screen "0004_Mixinghead" 1280x800, template "Navigation"
   on GenerateScreen: SetBit("DB704_MH_Value_Read"); SetBit("DB614_MH_State_Read"); SetTag("Navigation_7", 4); "MH_TestshotVisibility"()
   Button "Button_17" at 118,142 size 357x253; TextOff 'Text'
      Visibility <- "MH_Control_Visibility"
   TextField "Text field_43" at 173,150 size 158x29; Text 'Temperature'
      Visibility <- "MH_Control_Visibility"
   TextField "Text field_44" at 124,193 size 72x25; Text 'Actual:'
      Visibility <- "MH_Control_Visibility"
   TextField "Text field_45" at 124,226 size 100x25; Text 'Set value:'
      Visibility <- "MH_Control_Visibility"
   TextField "Text field_46" at 124,259 size 201x25; Text 'Warning upper limit:'
      Visibility <- "MH_Control_Visibility"
   TextField "Text field_47" at 124,292 size 199x25; Text 'Warning lower limit:'
      Visibility <- "MH_Control_Visibility"
   TextField "Text field_48" at 124,325 size 170x25; Text 'Fault upper limit:'
      Visibility <- "MH_Control_Visibility"
   TextField "Text field_49" at 124,358 size 168x25; Text 'Fault lower limit:'
      Visibility <- "MH_Control_Visibility"
   IOField "I/O field_29" at 336,189 size 81x32; FormatPattern 999.9
      Visibility <- "MH_Control_Visibility"
      ProcessValue <- "Temp_Actual"
   IOField "I/O field_30" at 336,222 size 81x32; Authorization "Operate"; FormatPattern 999.9
      Visibility <- "MH_Control_Visibility"
      ProcessValue <- "Temp_SetValue"
   IOField "I/O field_31" at 336,255 size 81x32; Authorization "Operate"; FormatPattern 999.9
      Visibility <- "MH_Control_Visibility"
      ProcessValue <- "Temp_Warning_Upper_Limit"
   IOField "I/O field_32" at 336,288 size 81x32; Authorization "Operate"; FormatPattern 999.9
      Visibility <- "MH_Control_Visibility"
      ProcessValue <- "Temp_Warning_Llower_Limit"
   IOField "I/O field_33" at 336,321 size 81x32; Authorization "Operate"; FormatPattern 999.9
      Visibility <- "MH_Control_Visibility"
      ProcessValue <- "Temp_Fault_Upper_Limit"
   IOField "I/O field_34" at 336,354 size 81x32; Authorization "Operate"; FormatPattern 999.9
      Visibility <- "MH_Control_Visibility"
      ProcessValue <- "Temp_Fault_Lower_Limit"
   Button "Button_18" at 417,148 size 51x41; TextOff 'Text'; PictureOff "images (1)"
      on Press: SetTag("MH_Control_Visibility", 0)
      Visibility <- "MH_Control_Visibility"
   TextField "Text field_78" at 424,193 size 46x25; Text 'ºC'
      Visibility <- "MH_Control_Visibility"
   IOField "I/O field_50" at 317,150 size 84x30; FormatPattern ????????????????????
      Visibility <- "MH_Control_Visibility"
      ProcessValue <- "Temp_Name"
   TextField "Text field_42" at 424,226 size 46x25; Text 'ºC'
      Visibility <- "MH_Control_Visibility"
   TextField "Text field_50" at 424,259 size 46x25; Text 'Δ ºC'
      Visibility <- "MH_Control_Visibility"
   TextField "Text field_51" at 424,292 size 46x25; Text 'Δ ºC'
      Visibility <- "MH_Control_Visibility"
   TextField "Text field_52" at 424,325 size 46x25; Text 'Δ ºC'
      Visibility <- "MH_Control_Visibility"
   TextField "Text field_53" at 424,358 size 46x25; Text 'Δ ºC'
      Visibility <- "MH_Control_Visibility"
   Button "Button_7" at 117,142 size 357x253; TextOff 'Text'
      Visibility <- "MH_Control_Visibility"
   TextField "Text field_92" at 216,154 size 160x29; Text 'Inerting Data'
      Visibility <- "MH_Control_Visibility"
   TextField "Text field_93" at 123,189 size 118x25; Text 'Ready time:'
      Visibility <- "MH_Control_Visibility"
   TextField "Text field_94" at 123,217 size 188x25; Text 'Max. Inerting time:'
      Visibility <- "MH_Control_Visibility"
   TextField "Text field_95" at 123,245 size 198x25; Text 'Limit value inerting:'
      Visibility <- "MH_Control_Visibility"
   TextField "Text field_96" at 123,273 size 121x25; Text 'Start filling:'
      Visibility <- "MH_Control_Visibility"
   TextField "Text field_97" at 123,301 size 134x25; Text 'Filling factor:'
      Visibility <- "MH_Control_Visibility"
   TextField "Text field_98" at 123,329 size 122x25; Text 'Start offset:'
      Visibility <- "MH_Control_Visibility"
   IOField "I/O field_58" at 308,189 size 81x25; Authorization "Operate"; FormatPattern 99999
      Visibility <- "MH_Control_Visibility"
      ProcessValue <- "DB704_MH_Value_MH_Inerting{0}_Ready_Time_after_Inert"
   IOField "I/O field_59" at 308,217 size 81x25; Authorization "Operate"; FormatPattern 99999
      Visibility <- "MH_Control_Visibility"
      ProcessValue <- "DB704_MH_Value_MH_Inerting{0}_Max_Inerting_Time"
   IOField "I/O field_60" at 308,245 size 81x25; Authorization "User administration"; FormatPattern 9999.9
      Visibility <- "MH_Control_Visibility"
      ProcessValue <- "DB704_MH_Value_MH_Inerting{0}_Reference_Value_Inert"
   IOField "I/O field_61" at 308,273 size 81x25; Authorization "Operate"; FormatPattern 99999
      Visibility <- "MH_Control_Visibility"
      ProcessValue <- "DB704_MH_Value_MH_Inerting{0}_Foam_density"
   IOField "I/O field_62" at 308,301 size 81x25; Authorization "Operate"; FormatPattern 999.9
      Visibility <- "MH_Control_Visibility"
      ProcessValue <- "DB704_MH_Value_MH_Inerting{0}_Inerting_factor"
   IOField "I/O field_63" at 308,329 size 81x25; Authorization "Operate"; FormatPattern 999.9
      Visibility <- "MH_Control_Visibility"
      ProcessValue <- "DB704_MH_Value_MH_Inerting{0}_Start_Offset"
   Button "Button_9" at 416,148 size 51x41; TextOff 'Text'; PictureOff "images (1)"
      on Press: SetTag("MH_Control_Visibility", 0)
      Visibility <- "MH_Control_Visibility"
   IOField "I/O field_64" at 308,357 size 81x25; Authorization "Operate"; FormatPattern 999.9
      Visibility <- "MH_Control_Visibility"
      ProcessValue <- "DB704_MH_Value_MH_Inerting{0}_Leakage_Value"
   TextField "Text field_111" at 123,357 size 97x25; Text 'Min.level:'
      Visibility <- "MH_Control_Visibility"
   TextField "Text field_99" at 403,189 size 46x25; Text 's'
      Visibility <- "MH_Control_Visibility"
   TextField "Text field_100" at 403,217 size 46x25; Text 's'
      Visibility <- "MH_Control_Visibility"
   TextField "Text field_101" at 403,245 size 46x25; Text 'g'
      Visibility <- "MH_Control_Visibility"
   TextField "Text field_102" at 404,273 size 57x25; Text 'g/dm'
      Visibility <- "MH_Control_Visibility"
   TextField "Text field_103" at 452,269 size 36x18; Text '3'
      Visibility <- "MH_Control_Visibility"
   TextField "Text field_104" at 403,329 size 46x25; Text 'L'
      Visibility <- "MH_Control_Visibility"
   TextField "Text field_105" at 403,357 size 46x25; Text 'L'
      Visibility <- "MH_Control_Visibility"
   Button "Button_24" at 417,149 size 51x41; TextOff 'Text'; PictureOff "images (1)"
      on Press: SetTag("MH_Control_Visibility", 0)
      Visibility <- "MH_Control_Visibility"
   Button "Button_25" at 118,143 size 357x253; TextOff 'Text'
      Visibility <- "MH_Control_Visibility"
   TextField "Text field_137" at 249,155 size 96x29; Text 'Blowing'
      Visibility <- "MH_Control_Visibility"
   TextField "Text field_138" at 124,215 size 137x25; Text 'Blowing time:'
      Visibility <- "MH_Control_Visibility"
   TextField "Text field_139" at 124,248 size 237x25; Text 'Blowing time after shot:'
      Visibility <- "MH_Control_Visibility"
   IOField "I/O field_79" at 346,215 size 81x25; Authorization "Operate"; FormatPattern 99999
      Visibility <- "MH_Control_Visibility"
      ProcessValue <- "DB704_MH_Value_MH_Inerting{0}_Purge_time"
   IOField "I/O field_80" at 346,248 size 81x25; Authorization "Operate"; FormatPattern 99999
      Visibility <- "MH_Control_Visibility"
      ProcessValue <- "DB704_MH_Value_MH_Inerting{0}_Purge_after_Shot"
   Button "Button_26" at 417,149 size 51x41; TextOff 'Text'; PictureOff "images (1)"
      on Press: SetTag("MH_Control_Visibility", 0)
      Visibility <- "MH_Control_Visibility"
   TextField "Text field_145" at 442,215 size 46x25; Text 's'
      Visibility <- "MH_Control_Visibility"
   TextField "Text field_146" at 442,248 size 46x25; Text 's'
      Visibility <- "MH_Control_Visibility"
   Button "spare_2" at 335,709 size 36x32; TextOff 'Text'
      Visibility <- "DB704_MH_Value_Mixinghead{0}_MH_Connection{1}_WithNozzle"
   Button "spare_3" at 335,748 size 36x32; TextOff 'Text'
      Visibility <- "DB704_MH_Value_Mixinghead{0}_MH_Connection{1}_WithNozzle"
   Button "spare_1" at 335,670 size 36x32; TextOff 'Text'
      Visibility <- "DB704_MH_Value_Mixinghead{0}_MH_Connection{1}_WithNozzle"
   Button "spare_10" at 473,748 size 36x32; TextOff 'Text'
      Visibility <- "DB704_MH_Value_Mixinghead{0}_MH_Connection{2}_WithNozzle"
   Button "spare_9" at 473,709 size 36x32; TextOff 'Text'
      Visibility <- "DB704_MH_Value_Mixinghead{0}_MH_Connection{2}_WithNozzle"
   Button "spare_4" at 473,670 size 36x32; TextOff 'Text'
      Visibility <- "DB704_MH_Value_Mixinghead{0}_MH_Connection{2}_WithNozzle"
   Button "spare_5" at 611,670 size 36x32; TextOff 'Text'
      Visibility <- "DB704_MH_Value_Mixinghead{0}_MH_Connection{3}_WithNozzle"
   Button "spare_11" at 611,709 size 36x32; TextOff 'Text'
      Visibility <- "DB704_MH_Value_Mixinghead{0}_MH_Connection{3}_WithNozzle"
   Button "spare_12" at 611,748 size 36x32; TextOff 'Text'
      Visibility <- "DB704_MH_Value_Mixinghead{0}_MH_Connection{3}_WithNozzle"
   Button "spare_14" at 749,748 size 36x32; TextOff 'Text'
      Visibility <- "DB704_MH_Value_Mixinghead{0}_MH_Connection{4}_WithNozzle"
   Button "spare_13" at 749,709 size 36x32; TextOff 'Text'
      Visibility <- "DB704_MH_Value_Mixinghead{0}_MH_Connection{4}_WithNozzle"
   Button "spare_6" at 749,670 size 36x32; TextOff 'Text'
      Visibility <- "DB704_MH_Value_Mixinghead{0}_MH_Connection{4}_WithNozzle"
   Button "spare_7" at 887,670 size 36x32; TextOff 'Text'
      Visibility <- "DB704_MH_Value_Mixinghead{0}_MH_Connection{5}_WithNozzle"
   Button "spare_15" at 887,709 size 36x32; TextOff 'Text'
      Visibility <- "DB704_MH_Value_Mixinghead{0}_MH_Connection{5}_WithNozzle"
   Button "spare_16" at 887,748 size 36x32; TextOff 'Text'
      Visibility <- "DB704_MH_Value_Mixinghead{0}_MH_Connection{5}_WithNozzle"
   Button "spare_17" at 1025,709 size 36x32; TextOff 'Text'
      Visibility <- "DB704_MH_Value_Mixinghead{0}_MH_Connection{6}_WithNozzle"
   Button "spare_18" at 1025,748 size 36x32; TextOff 'Text'
      Visibility <- "DB704_MH_Value_Mixinghead{0}_MH_Connection{6}_WithNozzle"
   Button "spare_8" at 1025,670 size 36x32; TextOff 'Text'
      Visibility <- "DB704_MH_Value_Mixinghead{0}_MH_Connection{6}_WithNozzle"
   Rectangle "Rectangle_43" at 746,666 size 138x40
      Visibility <- "DB614_MH_State_MH_Status{0}_QPB_Values_selected"
   Rectangle "Rectangle_40" at 470,627 size 138x40
      Visibility <- "DB614_MH_State_MH_Status{0}_QPB_Values_selected"
   Rectangle "Rectangle_35" at 608,627 size 138x40
      Visibility <- "DB614_MH_State_MH_Status{0}_QPB_Values_selected"
   Rectangle "Rectangle_36" at 746,627 size 138x40
      Visibility <- "DB614_MH_State_MH_Status{0}_QPB_Values_selected"
   Rectangle "Rectangle_37" at 884,627 size 138x40
      Visibility <- "DB614_MH_State_MH_Status{0}_QPB_Values_selected"
   Rectangle "Rectangle_38" at 1022,627 size 138x40
      Visibility <- "DB614_MH_State_MH_Status{0}_QPB_Values_selected"
   Rectangle "Rectangle_41" at 470,666 size 138x40
      Visibility <- "DB614_MH_State_MH_Status{0}_QPB_Values_selected"
   Rectangle "Rectangle_42" at 608,666 size 138x40
      Visibility <- "DB614_MH_State_MH_Status{0}_QPB_Values_selected"
   Rectangle "Rectangle_44" at 884,666 size 138x40
      Visibility <- "DB614_MH_State_MH_Status{0}_QPB_Values_selected"
   Rectangle "Rectangle_45" at 1022,666 size 138x40
      Visibility <- "DB614_MH_State_MH_Status{0}_QPB_Values_selected"
   Rectangle "Rectangle_46" at 470,705 size 138x40
      Visibility <- "DB614_MH_State_MH_Status{0}_QPB_Values_selected"
   Rectangle "Rectangle_47" at 608,705 size 138x40
      Visibility <- "DB614_MH_State_MH_Status{0}_QPB_Values_selected"
   Rectangle "Rectangle_48" at 746,705 size 138x40
      Visibility <- "DB614_MH_State_MH_Status{0}_QPB_Values_selected"
   Rectangle "Rectangle_49" at 884,705 size 138x40
      Visibility <- "DB614_MH_State_MH_Status{0}_QPB_Values_selected"
   Rectangle "Rectangle_50" at 1022,705 size 138x40
      Visibility <- "DB614_MH_State_MH_Status{0}_QPB_Values_selected"
   Rectangle "Rectangle_39" at 332,627 size 138x40
      Visibility <- "DB614_MH_State_MH_Status{0}_QPB_Values_selected"
   Rectangle "Rectangle_34" at 332,666 size 138x40
      Visibility <- "DB614_MH_State_MH_Status{0}_QPB_Values_selected"
   Rectangle "Rectangle_33" at 332,705 size 138x40
      Visibility <- "DB614_MH_State_MH_Status{0}_QPB_Values_selected"
   Button "Button_13" at 120,144 size 357x253; TextOff 'Text'
      Visibility <- "MH_Control_Visibility"
   TextField "Text field_6" at 177,156 size 111x29; Text 'Pressure'
      Visibility <- "MH_Control_Visibility"
   TextField "Text field_7" at 126,195 size 72x25; Text 'Actual:'
      Visibility <- "MH_Control_Visibility"
   TextField "Text field_8" at 126,228 size 100x25; Text 'Set value:'
      Visibility <- "MH_Control_Visibility"
   TextField "Text field_9" at 126,261 size 201x25; Text 'Warning upper limit:'
      Visibility <- "MH_Control_Visibility"
   TextField "Text field_19" at 126,294 size 199x25; Text 'Warning lower limit:'
      Visibility <- "MH_Control_Visibility"
   TextField "Text field_20" at 126,327 size 170x25; Text 'Fault upper limit:'
      Visibility <- "MH_Control_Visibility"
   TextField "Text field_21" at 126,360 size 168x25; Text 'Fault lower limit:'
      Visibility <- "MH_Control_Visibility"
   IOField "I/O field_12" at 311,192 size 81x32; Authorization "User administration"; FormatPattern 999.9
      Visibility <- "MH_Control_Visibility"
      ProcessValue <- "Press_Actual"
   IOField "I/O field_13" at 311,225 size 81x32; Authorization "Operate"; FormatPattern 999.9
      Visibility <- "MH_Control_Visibility"
      ProcessValue <- "Press_SetValue"
   IOField "I/O field_14" at 311,258 size 81x32; Authorization "Operate"; FormatPattern 999.9
      Visibility <- "MH_Control_Visibility"
      ProcessValue <- "Press_Warning_Upper_Limit"
   IOField "I/O field_15" at 311,291 size 81x32; Authorization "Operate"; FormatPattern 999.9
      Visibility <- "MH_Control_Visibility"
      ProcessValue <- "Press_Warning_Lower_Limit"
   IOField "I/O field_21" at 311,324 size 81x32; Authorization "Operate"; FormatPattern 999.9
      Visibility <- "MH_Control_Visibility"
      ProcessValue <- "Press_Fault_Upper_Limit"
   IOField "I/O field_22" at 311,357 size 81x32; Authorization "Operate"; FormatPattern 999.9
      Visibility <- "MH_Control_Visibility"
      ProcessValue <- "Press_Fault_Lower_Limit"
   TextField "Text field_22" at 417,195 size 46x25; Text 'bar'
      Visibility <- "MH_Control_Visibility"
   TextField "Text field_23" at 417,228 size 46x25; Text 'bar'
      Visibility <- "MH_Control_Visibility"
   TextField "Text field_24" at 417,261 size 55x25; Text 'Δ bar'
      Visibility <- "MH_Control_Visibility"
   TextField "Text field_25" at 417,294 size 55x25; Text 'Δ bar'
      Visibility <- "MH_Control_Visibility"
   TextField "Text field_26" at 417,327 size 55x25; Text 'Δ bar'
      Visibility <- "MH_Control_Visibility"
   TextField "Text field_27" at 417,360 size 55x25; Text 'Δ bar'
      Visibility <- "MH_Control_Visibility"
   Button "Button_14" at 419,150 size 51x41; TextOff 'Text'; PictureOff "images (1)"
      on Press: SetTag("MH_Control_Visibility", 0)
      Visibility <- "MH_Control_Visibility"
   TextField "Text field_28" at 417,195 size 46x25; Text 'bar'
      Visibility <- "MH_Control_Visibility"
   TextField "Text field_82" at 105,674 size 174x25; Text 'Pressure built up:'
      Visibility <- "DB614_MH_State_MH_Status{0}_QPB_Values_selected"
   TextField "Text field_83" at 105,710 size 146x25; Text 'Until pressure:'
      Visibility <- "DB614_MH_State_MH_Status{0}_QPB_Values_selected"
   TextField "Text field_85" at 277,673 size 46x25; Text 'g/s'
      Visibility <- "DB614_MH_State_MH_Status{0}_QPB_Values_selected"
   TextField "Text field_86" at 277,711 size 46x25; Text 'bar'
      Visibility <- "DB614_MH_State_MH_Status{0}_QPB_Values_selected"
   IOField "I/O field_41" at 370,631 size 94x32; FormatPattern 9999.99
      Visibility <- "DB614_MH_State_MH_Status{0}_QPB_Values_selected"
      ProcessValue <- "DB614_MH_State_MH_Connection{0}_ActFlow{1}"
   IOField "I/O field_42" at 370,669 size 94x32; Authorization "Operate"; FormatPattern 9999.99
      ProcessValue <- "DB704_MH_Value_Mixinghead{0}_MH_Connection{1}_FlowQPB"
      Visibility <- "DB614_MH_State_MH_Status{0}_QPB_Values_selected"
   IOField "I/O field_43" at 370,708 size 94x32; Authorization "Operate"; FormatPattern 9999.99
      ProcessValue <- "DB704_MH_Value_Mixinghead{0}_MH_Connection{1}_PressureQPB"
      Visibility <- "DB614_MH_State_MH_Status{0}_QPB_Values_selected"
   IOField "I/O field_44" at 508,631 size 94x32; FormatPattern 9999.99
      Visibility <- "DB614_MH_State_MH_Status{0}_QPB_Values_selected"
      ProcessValue <- "DB614_MH_State_MH_Connection{0}_ActFlow{2}"
   IOField "I/O field_45" at 508,670 size 94x32; Authorization "Operate"; FormatPattern 9999.99
      ProcessValue <- "DB704_MH_Value_Mixinghead{0}_MH_Connection{2}_FlowQPB"
      Visibility <- "DB614_MH_State_MH_Status{0}_QPB_Values_selected"
   IOField "I/O field_46" at 508,708 size 94x32; Authorization "Operate"; FormatPattern 9999.99
      ProcessValue <- "DB704_MH_Value_Mixinghead{0}_MH_Connection{2}_PressureQPB"
      Visibility <- "DB614_MH_State_MH_Status{0}_QPB_Values_selected"
   IOField "I/O field_49" at 278,156 size 84x30; Authorization "Operate"; FormatPattern ????????????????????
      Visibility <- "MH_Control_Visibility"
      ProcessValue <- "Press_Name"
   IOField "I/O field_109" at 646,631 size 94x32; FormatPattern 9999.99
      Visibility <- "DB614_MH_State_MH_Status{0}_QPB_Values_selected"
      ProcessValue <- "DB614_MH_State_MH_Connection{0}_ActFlow{3}"
   IOField "I/O field_110" at 646,670 size 94x32; Authorization "Operate"; FormatPattern 9999.99
      ProcessValue <- "DB704_MH_Value_Mixinghead{0}_MH_Connection{3}_FlowQPB"
      Visibility <- "DB614_MH_State_MH_Status{0}_QPB_Values_selected"
   IOField "I/O field_111" at 646,708 size 94x32; Authorization "Operate"; FormatPattern 9999.99
      ProcessValue <- "DB704_MH_Value_Mixinghead{0}_MH_Connection{3}_PressureQPB"
      Visibility <- "DB614_MH_State_MH_Status{0}_QPB_Values_selected"
   IOField "I/O field_112" at 784,631 size 94x32; FormatPattern 9999.99
      Visibility <- "DB614_MH_State_MH_Status{0}_QPB_Values_selected"
      ProcessValue <- "DB614_MH_State_MH_Connection{0}_ActFlow{4}"
   IOField "I/O field_113" at 784,670 size 94x32; Authorization "User administration"; FormatPattern 9999.99
      ProcessValue <- "DB704_MH_Value_Mixinghead{0}_MH_Connection{4}_FlowQPB"
      Visibility <- "DB614_MH_State_MH_Status{0}_QPB_Values_selected"
   IOField "I/O field_114" at 784,708 size 94x32; Authorization "Operate"; FormatPattern 9999.99
      ProcessValue <- "DB704_MH_Value_Mixinghead{0}_MH_Connection{4}_PressureQPB"
      Visibility <- "DB614_MH_State_MH_Status{0}_QPB_Values_selected"
   IOField "I/O field_115" at 922,631 size 94x32; FormatPattern 9999.99
      Visibility <- "DB614_MH_State_MH_Status{0}_QPB_Values_selected"
      ProcessValue <- "DB614_MH_State_MH_Connection{0}_ActFlow{5}"
   IOField "I/O field_116" at 922,670 size 94x32; Authorization "User administration"; FormatPattern 9999.99
      ProcessValue <- "DB704_MH_Value_Mixinghead{0}_MH_Connection{5}_FlowQPB"
      Visibility <- "DB614_MH_State_MH_Status{0}_QPB_Values_selected"
   IOField "I/O field_117" at 922,708 size 94x32; Authorization "User administration"; FormatPattern 9999.99
      ProcessValue <- "DB704_MH_Value_Mixinghead{0}_MH_Connection{5}_PressureQPB"
      Visibility <- "DB614_MH_State_MH_Status{0}_QPB_Values_selected"
   IOField "I/O field_118" at 1060,631 size 94x32; FormatPattern 9999.99
      Visibility <- "DB614_MH_State_MH_Status{0}_QPB_Values_selected"
      ProcessValue <- "DB614_MH_State_MH_Connection{0}_ActFlow{6}"
   IOField "I/O field_119" at 1060,670 size 94x32; Authorization "Operate"; FormatPattern 9999.99
      ProcessValue <- "DB704_MH_Value_Mixinghead{0}_MH_Connection{6}_FlowQPB"
      Visibility <- "DB614_MH_State_MH_Status{0}_QPB_Values_selected"
   IOField "I/O field_120" at 1060,708 size 94x32; Authorization "Operate"; FormatPattern 9999.99
      ProcessValue <- "DB704_MH_Value_Mixinghead{0}_MH_Connection{6}_PressureQPB"
      Visibility <- "DB614_MH_State_MH_Status{0}_QPB_Values_selected"
   Rectangle "Rectangle_51" at 608,744 size 138x40
      Visibility <- "DB614_MH_State_MH_Status{0}_QPB_Values_selected"
   Rectangle "Rectangle_52" at 746,744 size 138x40
      Visibility <- "DB614_MH_State_MH_Status{0}_QPB_Values_selected"
   Rectangle "Rectangle_53" at 884,744 size 138x40
      Visibility <- "DB614_MH_State_MH_Status{0}_QPB_Values_selected"
   Rectangle "Rectangle_54" at 1022,744 size 138x40
      Visibility <- "DB614_MH_State_MH_Status{0}_QPB_Values_selected"
   Rectangle "Rectangle_31" at 470,744 size 138x40
      Visibility <- "DB614_MH_State_MH_Status{0}_QPB_Values_selected"
   Rectangle "Rectangle_32" at 332,744 size 138x40
      Visibility <- "DB614_MH_State_MH_Status{0}_QPB_Values_selected"
   IOField "I/O field_5" at 371,631 size 94x32; FormatPattern 9999.99
      Visibility <- "DB614_MH_State_MH_Status{0}_QPB_Values_selected"
      ProcessValue <- "DB614_MH_State_MH_Connection{0}_ActFlow{1}"
   IOField "I/O field_6" at 371,669 size 94x32; Authorization "Operate"; FormatPattern 9999.99
      ProcessValue <- "DB704_MH_Value_Mixinghead{0}_MH_Connection{1}_Flow_red_Circ"
      Visibility <- "DB614_MH_State_MH_Status{0}_QPB_Values_selected"
   IOField "I/O field_7" at 371,708 size 94x32; Authorization "Operate"; FormatPattern 9999.99
      ProcessValue <- "DB704_MH_Value_Mixinghead{0}_MH_Connection{1}_Flow_HP_Circ"
      Visibility <- "DB614_MH_State_MH_Status{0}_QPB_Values_selected"
   IOField "I/O field_8" at 371,748 size 94x32; Authorization "Operate"; FormatPattern 9999.99
      ProcessValue <- "DB704_MH_Value_Mixinghead{0}_MH_Connection{1}_Flow_LP_Circ"
      Visibility <- "DB614_MH_State_MH_Status{0}_QPB_Values_selected"
   IOField "I/O field_11" at 509,748 size 92x32; Authorization "Operate"; FormatPattern 9999.99
      ProcessValue <- "DB704_MH_Value_Mixinghead{0}_MH_Connection{2}_Flow_LP_Circ"
      Visibility <- "DB614_MH_State_MH_Status{0}_QPB_Values_selected"
   IOField "I/O field_10" at 509,708 size 92x32; Authorization "Operate"; FormatPattern 9999.99
      ProcessValue <- "DB704_MH_Value_Mixinghead{0}_MH_Connection{2}_Flow_HP_Circ"
      Visibility <- "DB614_MH_State_MH_Status{0}_QPB_Values_selected"
   IOField "I/O field_9" at 509,670 size 92x32; Authorization "Operate"; FormatPattern 9999.99
      ProcessValue <- "DB704_MH_Value_Mixinghead{0}_MH_Connection{2}_Flow_red_Circ"
      Visibility <- "DB614_MH_State_MH_Status{0}_QPB_Values_selected"
   IOField "I/O field_4" at 509,631 size 92x32; FormatPattern 9999.99
      Visibility <- "DB614_MH_State_MH_Status{0}_QPB_Values_selected"
      ProcessValue <- "DB614_MH_State_MH_Connection{0}_ActFlow{2}"
   IOField "I/O field_92" at 647,631 size 92x32; FormatPattern 9999.99
      Visibility <- "DB614_MH_State_MH_Status{0}_QPB_Values_selected"
      ProcessValue <- "DB614_MH_State_MH_Connection{0}_ActFlow{3}"
   IOField "I/O field_93" at 647,670 size 92x32; Authorization "Operate"; FormatPattern 9999.99
      ProcessValue <- "DB704_MH_Value_Mixinghead{0}_MH_Connection{3}_Flow_red_Circ"
      Visibility <- "DB614_MH_State_MH_Status{0}_QPB_Values_selected"
   IOField "I/O field_94" at 647,708 size 92x32; Authorization "Operate"; FormatPattern 9999.99
      Visibility <- "DB614_MH_State_MH_Status{0}_QPB_Values_selected"
      ProcessValue <- "DB704_MH_Value_Mixinghead{0}_MH_Connection{3}_Flow_HP_Circ"
   IOField "I/O field_95" at 647,748 size 92x32; Authorization "Operate"; FormatPattern 9999.99
      ProcessValue <- "DB704_MH_Value_Mixinghead{0}_MH_Connection{3}_Flow_LP_Circ"
      Visibility <- "DB614_MH_State_MH_Status{0}_QPB_Values_selected"
   IOField "I/O Actual flow Con 4" at 785,631 size 92x32; FormatPattern 9999.99
      Visibility <- "DB614_MH_State_MH_Status{0}_QPB_Values_selected"
      ProcessValue <- "DB614_MH_State_MH_Connection{0}_ActFlow{4}"
   IOField "I/O field_96" at 785,670 size 92x32; Authorization "Operate"; FormatPattern 9999.99
      ProcessValue <- "DB704_MH_Value_Mixinghead{0}_MH_Connection{4}_Flow_red_Circ"
      Visibility <- "DB614_MH_State_MH_Status{0}_QPB_Values_selected"
   IOField "I/O field_98" at 785,748 size 92x32; Authorization "Operate"; FormatPattern 9999.99
      ProcessValue <- "DB704_MH_Value_Mixinghead{0}_MH_Connection{4}_Flow_LP_Circ"
      Visibility <- "DB614_MH_State_MH_Status{0}_QPB_Values_selected"
   IOField "I/O field_97" at 785,708 size 92x32; Authorization "Operate"; FormatPattern 9999.99
      ProcessValue <- "DB704_MH_Value_Mixinghead{0}_MH_Connection{4}_Flow_HP_Circ"
      Visibility <- "DB614_MH_State_MH_Status{0}_QPB_Values_selected"
   IOField "I/O field_102" at 923,631 size 92x32; FormatPattern 9999.99
      Visibility <- "DB614_MH_State_MH_Status{0}_QPB_Values_selected"
      ProcessValue <- "DB614_MH_State_MH_Connection{0}_ActFlow{5}"
   IOField "I/O field_103" at 923,670 size 92x32; Authorization "Operate"; FormatPattern 9999.99
      ProcessValue <- "DB704_MH_Value_Mixinghead{0}_MH_Connection{5}_Flow_red_Circ"
      Visibility <- "DB614_MH_State_MH_Status{0}_QPB_Values_selected"
   IOField "I/O field_104" at 923,708 size 92x32; Authorization "Operate"; FormatPattern 9999.99
      ProcessValue <- "DB704_MH_Value_Mixinghead{0}_MH_Connection{5}_Flow_HP_Circ"
      Visibility <- "DB614_MH_State_MH_Status{0}_QPB_Values_selected"
   IOField "I/O field_105" at 923,748 size 92x32; Authorization "Operate"; FormatPattern 9999.99
      ProcessValue <- "DB704_MH_Value_Mixinghead{0}_MH_Connection{5}_Flow_LP_Circ"
      Visibility <- "DB614_MH_State_MH_Status{0}_QPB_Values_selected"
   IOField "I/O field_108" at 1061,748 size 92x32; Authorization "Operate"; FormatPattern 9999.99
      ProcessValue <- "DB704_MH_Value_Mixinghead{0}_MH_Connection{6}_Flow_LP_Circ"
      Visibility <- "DB614_MH_State_MH_Status{0}_QPB_Values_selected"
   IOField "I/O field_107" at 1061,708 size 92x32; Authorization "Operate"; FormatPattern 9999.99
      ProcessValue <- "DB704_MH_Value_Mixinghead{0}_MH_Connection{6}_Flow_HP_Circ"
      Visibility <- "DB614_MH_State_MH_Status{0}_QPB_Values_selected"
   IOField "I/O field_106" at 1061,670 size 92x32; Authorization "Operate"; FormatPattern 9999.99
      ProcessValue <- "DB704_MH_Value_Mixinghead{0}_MH_Connection{6}_Flow_red_Circ"
      Visibility <- "DB614_MH_State_MH_Status{0}_QPB_Values_selected"
   IOField "I/O field_101" at 1061,631 size 92x32; FormatPattern 9999.99
      Visibility <- "DB614_MH_State_MH_Status{0}_QPB_Values_selected"
      ProcessValue <- "DB614_MH_State_MH_Connection{0}_ActFlow{6}"
   Rectangle "Rectangle_69" at 333,745 size 136x38
      Visibility <- "DB704_MH_Value_Mixinghead{0}_WithLPCirculation"
   Rectangle "Rectangle_70" at 471,745 size 136x38
      Visibility <- "DB704_MH_Value_Mixinghead{0}_WithLPCirculation"
   Rectangle "Rectangle_71" at 609,745 size 136x38
      Visibility <- "DB704_MH_Value_Mixinghead{0}_WithLPCirculation"
   Rectangle "Rectangle_72" at 747,745 size 136x38
      Visibility <- "DB704_MH_Value_Mixinghead{0}_WithLPCirculation"
   Rectangle "Rectangle_73" at 885,745 size 136x38
      Visibility <- "DB704_MH_Value_Mixinghead{0}_WithLPCirculation"
   Rectangle "Rectangle_74" at 1023,745 size 136x38
      Visibility <- "DB704_MH_Value_Mixinghead{0}_WithLPCirculation"
   Rectangle "Rectangle_68" at 104,745 size 227x38
      Visibility <- "DB704_MH_Value_Mixinghead{0}_WithLPCirculation"
   Button "Template_Button_41" at 16,724 size 68x66; TextOff 'Text'; PictureList "Ico_navigation_2"; PictureOff "Setting_Nav_7"; Authorization "User administration"
      on Click: ActivateScreen("0005_Mixinghead Settting", 0)
      ProcessValue <- "Nav_7"
      Visibility <- "NavUserChange"
   Rectangle "Rectangle_55" at 332,625 size 138x167
      Visibility <- "DB704_MH_Value_Mixinghead{0}_AmountComponent"
   Rectangle "Rectangle_56" at 470,625 size 138x167
      Visibility <- "DB704_MH_Value_Mixinghead{0}_AmountComponent"
   Rectangle "Rectangle_57" at 608,625 size 138x167
      Visibility <- "DB704_MH_Value_Mixinghead{0}_AmountComponent"
   Rectangle "Rectangle_58" at 746,625 size 138x167
      Visibility <- "DB704_MH_Value_Mixinghead{0}_AmountComponent"
   Rectangle "Rectangle_59" at 884,625 size 138x167
      Visibility <- "DB704_MH_Value_Mixinghead{0}_AmountComponent"
   Rectangle "Rectangle_60" at 1022,625 size 138x167
      Visibility <- "DB704_MH_Value_Mixinghead{0}_AmountComponent"
   TextField "Text field_34" at 768,446 size 94x25; Text 'ºC'
      Visibility <- "DB704_MH_Value_Mixinghead{0}_AmountComponent"
   TextField "Text field_35" at 768,421 size 94x25; Text 'bar'
      Visibility <- "DB704_MH_Value_Mixinghead{0}_AmountComponent"
   TextField "Text field_36" at 768,473 size 94x25; Text 'bar'
      Visibility <- "DB704_MH_Value_Mixinghead{0}_AmountComponent"
   TextField "Text field_37" at 768,527 size 94x25; Text 'bar'
      Visibility <- "DB704_MH_Value_Mixinghead{0}_AmountComponent"
   TextField "Text field_38" at 768,499 size 94x25; Text 'ºC'
      Visibility <- "DB704_MH_Value_Mixinghead{0}_AmountComponent"
   TextField "Text field_39" at 768,554 size 94x25; Text 'ºC'
      Visibility <- "DB704_MH_Value_Mixinghead{0}_AmountComponent"
   TextField "Text field_160" at 488,421 size 94x25; Text 'bar'
      Visibility <- "DB704_MH_Value_Mixinghead{0}_AmountComponent"
   TextField "Text field_29" at 488,447 size 94x25; Text 'ºC'
      Visibility <- "DB704_MH_Value_Mixinghead{0}_AmountComponent"
   TextField "Text field_30" at 488,473 size 94x25; Text 'bar'
      Visibility <- "DB704_MH_Value_Mixinghead{0}_AmountComponent"
   TextField "Text field_31" at 488,499 size 94x25; Text 'ºC'
      Visibility <- "DB704_MH_Value_Mixinghead{0}_AmountComponent"
   TextField "Text field_32" at 488,527 size 94x25; Text 'bar'
      Visibility <- "DB704_MH_Value_Mixinghead{0}_AmountComponent"
   TextField "Text field_33" at 488,554 size 94x25; Text 'ºC'
      Visibility <- "DB704_MH_Value_Mixinghead{0}_AmountComponent"
   Button "Button_1" at 485,144 size 395x266; TextOff 'Text'
      Visibility <- "DB704_MH_Value_Mixinghead{0}_WithCleaningPiston"
   IOField "I/O field_78" at 488,499 size 67x25; FormatPattern 999.9
      Visibility <- "DB704_MH_Value_Mixinghead{0}_AmountComponent"
      ProcessValue <- "DB604_PV_Mixinghead_Mixinghead{0}_Temperature_Connection{3}_PV_ActV_Value"
   IOField "I/O field_77" at 488,473 size 67x25; FormatPattern 999.9
      Visibility <- "DB704_MH_Value_Mixinghead{0}_AmountComponent"
      ProcessValue <- "DB604_PV_Mixinghead_Mixinghead{0}_Pressure_Connection{3}_PV_ActV_Value"
   IOField "I/O field_17" at 488,447 size 67x25; FormatPattern 999.9
      Visibility <- "DB704_MH_Value_Mixinghead{0}_AmountComponent"
      ProcessValue <- "DB604_PV_Mixinghead_Mixinghead{0}_Temperature_Connection{1}_PV_ActV_Value"
   IOField "I/O field_16" at 488,421 size 67x25; FormatPattern 999.9
      Visibility <- "DB704_MH_Value_Mixinghead{0}_AmountComponent"
      ProcessValue <- "DB604_PV_Mixinghead_Mixinghead{0}_Pressure_Connection{1}_PV_ActV_Value"
   GraphicView "Graphic view_9" at 593,536 size 32x28; Picture "man mode"
      Visibility <- "DB123_MH_IO_Signals_MH{0}_IN_MH_Manual_Mode"
   TextField "Text field_1" at 513,153 size 87x25; Text 'CP Back:'
      Visibility <- "DB704_MH_Value_Mixinghead{0}_WithCleaningPiston"
   TextField "Text field_2" at 513,183 size 167x25; Text 'CP Front Manual:'
      Visibility <- "DB704_MH_Value_Mixinghead{0}_WithCleaningPiston"
   TextField "Text field_3" at 513,213 size 194x25; Text 'CP Front automatic:'
      Visibility <- "DB704_MH_Value_Mixinghead{0}_WithCleaningPiston"
   Button "Button_11" at 904,142 size 81x116; TextOff 'Text'
      Visibility <- "DB704_MH_Value_Mixinghead{0}_Cleaning_Piston_Spare_19"
   Button "Button_12" at 987,141 size 81x116; TextOff 'Text'
   Button "b_QPB" at 122,551 size 54x54; TextOff 'Text'; PictureList "MH"
      ProcessValue <- "DB614_MH_State_MH_Status{0}_QPB_Values_selected"
      on Click: InvertBit("DB614_MH_State_MH_Status{0}_QPB_Values_selected")
   IOField "CP_Back" at 752,153 size 85x25; Authorization "Operate"; FormatPattern 99999
      ProcessValue <- "DB704_MH_Value_Mixinghead{0}_Cleaning_Piston_RestTimeBack"
      Visibility <- "DB704_MH_Value_Mixinghead{0}_WithCleaningPiston"
   IOField "I/O field_2" at 752,183 size 85x25; Authorization "Operate"; FormatPattern 99999
      ProcessValue <- "DB704_MH_Value_Mixinghead{0}_Cleaning_Piston_RestTimeFrontManual"
      Visibility <- "DB704_MH_Value_Mixinghead{0}_WithCleaningPiston"
   IOField "I/O field_3" at 752,213 size 85x25; Authorization "Operate"; FormatPattern 99999
      ProcessValue <- "DB704_MH_Value_Mixinghead{0}_Cleaning_Piston_RestTimeFront"
      Visibility <- "DB704_MH_Value_Mixinghead{0}_WithCleaningPiston"
   IOField "I/O field_20" at 696,536 size 32x28; FormatPattern 99
      ProcessValue <- "DB123_MH_IO_Signals_MH{0}_IN_MH_Prog_No_MH"
   IOField "I/O field_55" at 752,243 size 85x25; Authorization "Operate"; FormatPattern 99999
      Visibility <- "DB704_MH_Value_Mixinghead{0}_Cleaning_Piston_CP_withInterval"
      ProcessValue <- "DB704_MH_Value_Mixinghead{0}_Cleaning_Piston_IntervalCounts"
   IOField "I/O field_56" at 752,273 size 85x25; Authorization "Operate"; FormatPattern 99999
      Visibility <- "DB704_MH_Value_Mixinghead{0}_Cleaning_Piston_CP_withInterval"
      ProcessValue <- "DB704_MH_Value_Mixinghead{0}_Cleaning_Piston_IntervalRestTimeFront"
   TextField "Text field_87" at 513,243 size 118x25; Text 'CP Interval:'
      Visibility <- "DB704_MH_Value_Mixinghead{0}_Cleaning_Piston_CP_withInterval"
   TextField "Text field_88" at 513,273 size 172x25; Text 'CP Interval front:'
      Visibility <- "DB704_MH_Value_Mixinghead{0}_Cleaning_Piston_CP_withInterval"
   TextField "Text field_89" at 513,303 size 168x25; Text 'CP Interval back:'
      Visibility <- "DB704_MH_Value_Mixinghead{0}_Cleaning_Piston_CP_withInterval"
   IOField "I/O field_57" at 752,303 size 85x25; Authorization "Operate"; FormatPattern 99999
      Visibility <- "DB704_MH_Value_Mixinghead{0}_Cleaning_Piston_CP_withInterval"
      ProcessValue <- "DB704_MH_Value_Mixinghead{0}_Cleaning_Piston_IntervalRestTimeBack"
   TextField "Text field_90" at 513,338 size 90x25; Text 'Inerting:'
      Visibility <- "DB704_MH_Value_Mixinghead{0}_WithInerting"
   TextField "Text field_91" at 513,373 size 89x25; Text 'Blowing:'
      Visibility <- "DB704_MH_Value_Mixinghead{0}_WithMHVenting"
   Button "Button_2" at 823,335 size 45x30; TextOff 'Text'; PictureOff "obeng"
      Visibility <- "DB704_MH_Value_Mixinghead{0}_WithInerting"
      on Click: SetTag("MH_Control_Visibility", 5)
   Button "Button_4" at 824,370 size 45x30; TextOff 'Text'; PictureOff "obeng"
      Visibility <- "DB704_MH_Value_Mixinghead{0}_WithMHVenting"
      on Click: SetTag("MH_Control_Visibility", 6)
   Button "b_MH_Increase" at 789,95 size 46x32; TextOff 'Text'; PictureOff "right arrow"
      on Click: function_dd21b452("DB614_MH_State_ReadDeviceNo", 1)
   Button "b_MH_Decrease" at 267,95 size 46x32; TextOff 'Text'; PictureOff "left arrow"
      on Click: function_b9b71300("DB614_MH_State_ReadDeviceNo", 1)
      ObjectEnable <- "DB614_MH_State_ReadDeviceNo"
   Button "b_MH_name" at 326,95 size 451x32; TextOff 'MH 01'; TextList "MH_NO"
      ProcessValue <- "DB614_MH_State_ReadDeviceNo"
   Button "Button_27" at 1097,414 size 81x116; TextOff 'Text'
      Visibility <- "DB704_MH_Value_Mixinghead{0}_WithHeating"
   Button "Button_28" at 1014,414 size 81x116; TextOff 'Text'
      Visibility <- "DB704_MH_Value_Mixinghead{0}_WithHeating"
   Button "Button_29" at 223,495 size 81x116; TextOff 'Text'
      Visibility <- "DB704_MH_Value_Mixinghead{0}_WithInerting"
   Button "Button_15" at 1070,141 size 81x116; TextOff 'Text'
   Button "Button_16" at 107,430 size 94x25; TextOff 'N2 Set'
      Visibility <- "DB704_MH_Value_Mixinghead{0}_WithInerting"
   Button "Button_20" at 107,455 size 94x25; TextOff 'N2 actual'
      Visibility <- "DB704_MH_Value_Mixinghead{0}_WithInerting"
   GraphicView "Graphic view_3" at 626,423 size 104x112; Picture "images_4"
   IOField "I/O field_81" at 488,527 size 67x25; FormatPattern 999.9
      Visibility <- "DB704_MH_Value_Mixinghead{0}_AmountComponent"
      ProcessValue <- "DB604_PV_Mixinghead_Mixinghead{0}_Pressure_Connection{5}_PV_ActV_Value"
   IOField "I/O field_82" at 488,554 size 67x25; FormatPattern 999.9
      Visibility <- "DB704_MH_Value_Mixinghead{0}_AmountComponent"
      ProcessValue <- "DB604_PV_Mixinghead_Mixinghead{0}_Temperature_Connection{5}_PV_ActV_Value"
   IOField "I/O field_18" at 768,421 size 67x25; FormatPattern 999.9
      Visibility <- "DB704_MH_Value_Mixinghead{0}_AmountComponent"
      ProcessValue <- "DB604_PV_Mixinghead_Mixinghead{0}_Pressure_Connection{2}_PV_ActV_Value"
   IOField "I/O field_19" at 768,446 size 67x25; FormatPattern 999.9
      Visibility <- "DB704_MH_Value_Mixinghead{0}_AmountComponent"
      ProcessValue <- "DB604_PV_Mixinghead_Mixinghead{0}_Temperature_Connection{2}_PV_ActV_Value"
   IOField "I/O field_83" at 768,473 size 67x25; FormatPattern 999.9
      Visibility <- "DB704_MH_Value_Mixinghead{0}_AmountComponent"
      ProcessValue <- "DB604_PV_Mixinghead_Mixinghead{0}_Pressure_Connection{4}_PV_ActV_Value"
   IOField "I/O field_84" at 768,499 size 67x25; FormatPattern 999.9
      Visibility <- "DB704_MH_Value_Mixinghead{0}_AmountComponent"
      ProcessValue <- "DB604_PV_Mixinghead_Mixinghead{0}_Temperature_Connection{4}_PV_ActV_Value"
   IOField "I/O field_85" at 768,527 size 67x25; FormatPattern 999.9
      Visibility <- "DB704_MH_Value_Mixinghead{0}_AmountComponent"
      ProcessValue <- "DB604_PV_Mixinghead_Mixinghead{0}_Pressure_Connection{6}_PV_ActV_Value"
   IOField "I/O field_86" at 768,554 size 67x25; FormatPattern 999.9
      Visibility <- "DB704_MH_Value_Mixinghead{0}_AmountComponent"
      ProcessValue <- "DB604_PV_Mixinghead_Mixinghead{0}_Temperature_Connection{6}_PV_ActV_Value"
   TextField "Text field_5" at 838,213 size 46x25; Text 's'
      Visibility <- "DB704_MH_Value_Mixinghead{0}_WithCleaningPiston"
   TextField "Text field_4" at 838,180 size 46x25; Text 's'
      Visibility <- "DB704_MH_Value_Mixinghead{0}_WithCleaningPiston"
   TextField "Text field_15" at 838,151 size 46x25; Text 's'
      Visibility <- "DB704_MH_Value_Mixinghead{0}_WithCleaningPiston"
   GraphicView "Graphic view_1" at 921,208 size 48x40; Picture "Service"
      Visibility <- "DB704_MH_Value_Mixinghead{0}_Cleaning_Piston_Spare_19"
   GraphicView "Graphic view_2" at 1010,208 size 40x40; Picture "HP"
   GraphicView "Graphic view_4" at 238,564 size 48x40; Picture "Inerting"
      Visibility <- "DB704_MH_Value_Mixinghead{0}_WithInerting"
   GraphicIOField "Cleaning Piston Picture" at 1088,208 size 48x40; PictureList "CleaningPiston"
      ProcessValue <- "DB614_MH_State_MH_Status{0}_Switch_Service_ON_OFF"
   GraphicView "Graphic view_5" at 630,536 size 32x28; Picture "cp2"
      Visibility <- "DB614_MH_State_MH_Status{0}_Switch_Service_ON_OFF"
   GraphicView "Graphic view_6" at 1030,482 size 48x40; Picture "Refilling From barrel"
      Visibility <- "DB704_MH_Value_Mixinghead{0}_WithHeating"
   GraphicView "Graphic view_7" at 1111,482 size 48x40; Picture "refill_1"
      Visibility <- "DB704_MH_Value_Mixinghead{0}_WithHeating"
   Rectangle "Rectangle_61" at 996,149 size 64x56
      Appearance <- "DB614_MH_State_MH_Status{0}_State_HP"
   Rectangle "Rectangle_62" at 1079,149 size 64x56
      Appearance <- "DB614_MH_State_MH_Status{0}_State_Service"
   GraphicIOField "Graphic I/O field_2" at 1004,153 size 48x48; PictureList "mh_switch_HP"
      ProcessValue <- "tes_3"
   GraphicIOField "Graphic I/O field_3" at 1087,153 size 48x48; PictureList "ON_OFF_SWITCH"
      ProcessValue <- "DB614_MH_State_MH_Status{0}_Switch_Service_ON_OFF"
   Button "Button_41" at 1068,135 size 88x128; TextOff 'Text'
      on Click: InvertBit("DB614_MH_State_MH_Status{0}_Switch_Service_ON_OFF")
   Button "Button_42" at 984,135 size 88x128; TextOff 'Text'
      on Click: InvertBit("DB614_MH_State_MH_Status{0}_Switch_HP_ON_OFF")
   Rectangle "Rectangle_63" at 912,150 size 64x56
      Visibility <- "DB704_MH_Value_Mixinghead{0}_Cleaning_Piston_Spare_19"
      Appearance <- "HMI_Tag_1"
   GraphicIOField "Graphic I/O field_4" at 920,155 size 48x48; PictureList "ON_OFF_SWITCH"
      Visibility <- "DB704_MH_Value_Mixinghead{0}_Cleaning_Piston_Spare_19"
      ProcessValue <- "DB614_MH_State_MH_CleaningPiston{0}_Switch_CP_Forward"
   Rectangle "Rectangle_64" at 232,503 size 64x56
      Visibility <- "DB704_MH_Value_Mixinghead{0}_WithInerting"
      Appearance <- "DB704_MH_Value_MH_Inerting{0}_with_Purge"
   GraphicIOField "Graphic I/O field_5" at 240,508 size 48x48; PictureList "ON_OFF_SWITCH"
      Visibility <- "DB704_MH_Value_Mixinghead{0}_WithInerting"
      ProcessValue <- "DB704_MH_Value_MH_Inerting{0}_with_Purge"
   Button "Button_43" at 899,135 size 88x128; TextOff 'Text'
      on Click: InvertBit("DB614_MH_State_MH_CleaningPiston{0}_Switch_CP_Forward")
      Visibility <- "DB704_MH_Value_Mixinghead{0}_Cleaning_Piston_Spare_19"
   Rectangle "Rectangle_65" at 1023,422 size 64x56
      Visibility <- "DB704_MH_Value_Mixinghead{0}_WithHeating"
   GraphicIOField "Graphic I/O field_6" at 1031,427 size 48x48; PictureList "ON_OFF_SWITCH"
      Visibility <- "DB704_MH_Value_Mixinghead{0}_WithHeating"
      ProcessValue <- "tes_1"
   Button "Button_44" at 1010,410 size 88x128; TextOff 'Text'
      on Click: InvertBit("DB612_Tank_State_Tank{0}_Switch_Refilling_ON_OFF")
      Visibility <- "DB704_MH_Value_Mixinghead{0}_WithHeating"
   Rectangle "Rectangle_66" at 1105,422 size 64x56
      Visibility <- "DB704_MH_Value_Mixinghead{0}_WithHeating"
   GraphicIOField "Graphic I/O field_7" at 1113,427 size 48x48; PictureList "ON_OFF_SWITCH"
      Visibility <- "DB704_MH_Value_Mixinghead{0}_WithHeating"
      ProcessValue <- "tes_2"
   Button "Button_45" at 1095,410 size 88x128; TextOff 'Text'
      Visibility <- "DB704_MH_Value_Mixinghead{0}_WithHeating"
   Button "Button_46" at 219,488 size 88x128; TextOff 'Text'
      on Click: InvertBit("DB704_MH_Value_MH_Inerting{0}_with_Purge")
      Visibility <- "DB704_MH_Value_Mixinghead{0}_WithInerting"
   GraphicView "Alarm Indicator Pump2_1" at 658,467 size 25x25; Picture "AlarmState2"
      Visibility <- "DB614_MH_State_MH_Status{0}_FaultExist"
   Button "b_Pump2_1" at 644,456 size 56x48; TextOff 'Text'
      on Press: ActivateScreen("0024_ActualFaults", 0); SetTag("Alarm_Filter_Tag", 1); SetTag("NavScreenChange", 0)
      ObjectEnable <- "DB614_MH_State_MH_Status{0}_FaultExist"
   GraphicView "Graphic view_8" at 593,536 size 32x28; Picture "automatic mode"
      Visibility <- "DB123_MH_IO_Signals_MH{0}_IN_MH_Auto_Mode"
   Button "Button_3" at 987,271 size 81x116; TextOff 'Text'
      Visibility <- "DB614_MH_State_MH_Status{0}_Switch_Testshot_B_ON_OFF"
   GraphicIOField "Cleaning Piston Picture_1" at 1005,338 size 48x40; PictureList "Tesshot_A"
      ProcessValue <- "DB614_MH_State_MH_Status{0}_Switch_Testshot_A_ON_OFF"
      Visibility <- "DB614_MH_State_MH_Status{0}_Switch_Testshot_B_ON_OFF"
   Rectangle "Rectangle_1" at 996,279 size 64x56
      Appearance <- "DB614_MH_State_MH_Status{0}_State_Testshot_A"
      Visibility <- "DB614_MH_State_MH_Status{0}_Switch_Testshot_B_ON_OFF"
   GraphicIOField "Graphic I/O field_1" at 1004,283 size 48x48; PictureList "ON_OFF_SWITCH"
      ProcessValue <- "DB614_MH_State_MH_Status{0}_Switch_Testshot_A_ON_OFF"
      Visibility <- "DB614_MH_State_MH_Status{0}_Switch_Testshot_B_ON_OFF"
   Button "Button_21" at 985,265 size 88x128; TextOff 'Text'
      on Click: InvertBit("DB614_MH_State_MH_Status{0}_Switch_Testshot_A_ON_OFF")
      Visibility <- "DB614_MH_State_MH_Status{0}_Switch_Testshot_B_ON_OFF"
   Button "Button_22" at 1074,271 size 81x116; TextOff 'Text'
      Visibility <- "DB614_MH_State_MH_Status{0}_Switch_Testshot_A_ON_OFF"
   GraphicIOField "Cleaning Piston Picture_2" at 1092,338 size 48x40; PictureList "Tesshot_B"
      ProcessValue <- "DB614_MH_State_MH_Status{0}_Switch_Testshot_B_ON_OFF"
      Visibility <- "DB614_MH_State_MH_Status{0}_Switch_Testshot_A_ON_OFF"
   Rectangle "Rectangle_67" at 1083,279 size 64x56
      Appearance <- "DB614_MH_State_MH_Status{0}_State_Testshot_B"
      Visibility <- "DB614_MH_State_MH_Status{0}_Switch_Testshot_A_ON_OFF"
   GraphicIOField "Graphic I/O field_8" at 1091,283 size 48x48; PictureList "ON_OFF_SWITCH"
      ProcessValue <- "DB614_MH_State_MH_Status{0}_Switch_Testshot_B_ON_OFF"
      Visibility <- "DB614_MH_State_MH_Status{0}_Switch_Testshot_A_ON_OFF"
   Button "Button_39" at 1072,265 size 88x128; TextOff 'Text'
      on Click: InvertBit("DB614_MH_State_MH_Status{0}_Switch_Testshot_B_ON_OFF")
      Visibility <- "DB614_MH_State_MH_Status{0}_Switch_Testshot_A_ON_OFF"
   Button "Button_8" at 489,421 size 94x25; TextOff 'bar'
      on Press: SetTag("MH_Control_Visibility", 1); SetTag("Press_Control_Screen", 0)
      Visibility <- "DB704_MH_Value_Mixinghead{0}_AmountComponent"
   Button "Button_10" at 489,447 size 94x25; TextOff 'Text'
      on Press: SetTag("MH_Control_Visibility", 2); SetTag("Temp_Control_Screen", 0)
      Visibility <- "DB704_MH_Value_Mixinghead{0}_AmountComponent"
   Button "Button_30" at 489,473 size 94x25; TextOff 'bar'